// TIA Portal project "DistributoreCaffè" (V19)

(* hardware
DEVICE "S7-1200 station_1"  S7-1200 Station
   slot 0: "Telaio di montaggio_0"  S7-1200 Rack  Rack  V1.0
   slot 1: "PLC"  CPU 1212C DC/DC/Rly  6ES7 212-1HE40-0XB0  V4.6
DEVICE "HMI"  KTP900 Basic PN
   slot 0: "HMI_1"  KTP900 Basic PN  6AV2 123-2JB03-0AX0  17.0.0.0
   slot 1: "HMI_RT_1"  KTP900 Basic PN  6AV2 123-2JB03-0AX0  17.0.0.0
   slot 5: "HMI_1.IE_CP_1"  PROFINET Interface  17.0.0.0
      slot 1: "Interfaccia_1 PROFINET"  PROFINET Interface
         slot 1: "Porta_1"  Port
*)

// ===== PLC "PLC"  CPU 1212C DC/DC/Rly =====

TYPE "CreditoResto"
   STRUCT
      "5Cents" : Real;
      "10Cents" : Real;
      "20Cents" : Real;
      "50Cents" : Real;
      "1Euro" : Real;
      "2Euro" : Real;
   END_STRUCT;
END_TYPE

TYPE "RestoUtente"
   STRUCT
      "5Cents" : SInt;
      "10Cents" : SInt;
      "20Cents" : SInt;
      "50Cents" : SInt;
      "1Euro" : SInt;
      "2Euro" : SInt;
   END_STRUCT;
END_TYPE

TYPE "Prezzo"
   STRUCT
      Bevanda : String;
      Prezzo : Real;
   END_STRUCT;
END_TYPE

DATA_BLOCK "HMI"   // DB1
{ S7_Optimized_Access := 'TRUE' }
VERSION : 0.1
   VAR
      I5cents : Bool;
      I10Cents : Bool;
      I20Cents : Bool;
      I50Cents : Bool;
      I1Euro : Bool;
      I2Euro : Bool;
   END_VAR
   VAR RETAIN
      Resto : "RestoUtente";
   END_VAR
   VAR
      ValvolaBicchiere : Bool;
      ValvolaPaletta : Bool;
      ValvolaCaffè : Bool;
      ValvolaLatte : Bool;
      ValvolaGrappa : Bool;
      ValvolaZucchero : Bool;
      PrelievoProdotto : Bool;
   END_VAR
   VAR RETAIN
      ProdottoPronto : Bool;
   END_VAR
   VAR
      Corto : Bool;
      CortoMacchiato : Bool;
      CortoCorretto : Bool;
      CortoMacchiatoCorretto : Bool;
      Lungo : Bool;
      LungoMacchiato : Bool;
      LungoCorretto : Bool;
      LungoMacchiatoCorretto : Bool;
      ConfermaOrdine : Bool;
      BicchieriScarico : Bool;
      PaletteScarico : Bool;
      CaffèScarico : Bool;
      LatteScarico : Bool;
      GrappaScarico : Bool;
      ZuccheroScarico : Bool;
      Bicchieri : Int;
      Palette : Int;
      Caffè : SInt;
      Latte : SInt;
      Grappa : SInt;
      Zucchero : SInt;
      Credito : Real;
      Introiti : Real;
      PrelievoIntroiti : Bool;
      CreditoInsufficiente : Bool;
      QuantitàZuccheroSelezionata : SInt;
      RiduzioneZucchero : Bool;
      IncrementoZucchero : Bool;
      ProdottoInPreparazione : Bool;
   END_VAR
BEGIN
END_DATA_BLOCK

DATA_BLOCK "Sistema"   // DB2
{ S7_Optimized_Access := 'TRUE' }
VERSION : 0.1
   VAR RETAIN
      CreditoResto : "CreditoResto";
   END_VAR
   VAR
      PConfermaOrdine : Bool;
      BloccoInterfacciaUtente : Bool;
      NPrelievoProdotto : Bool;
      BevandaSelezionata : SInt;
      PCorto : Bool;
      PCortoMacchiato : Bool;
      PCortoCorretto : Bool;
      PCortoMacchiatoCorretto : Bool;
      PLungo : Bool;
      PLungoMacchiato : Bool;
      PLungoCorretto : Bool;
      PLungoMacchiatoCorretto : Bool;
      PPiùZucchero : Bool;
      PMenoZucchero : Bool;
   END_VAR
   VAR RETAIN
      Prezzi : Array[1..8] of "Prezzo";
   END_VAR
   VAR
      PBloccoInterfacciaUtente : Bool;
      NPrelievoProdotto2 : Bool;
   END_VAR
BEGIN
   CreditoResto."5Cents" := 5.0;
   CreditoResto."10Cents" := 5.0;
   CreditoResto."20Cents" := 5.0;
   CreditoResto."50Cents" := 5.0;
   CreditoResto."1Euro" := 5.0;
   CreditoResto."2Euro" := 5.0;
   Prezzi[1].Bevanda := 'Corto';
   Prezzi[1].Prezzo := 0.3;
   Prezzi[2].Bevanda := 'CortoMacchiato';
   Prezzi[2].Prezzo := 0.4;
   Prezzi[3].Bevanda := 'CortoCorretto';
   Prezzi[3].Prezzo := 0.4;
   Prezzi[4].Bevanda := 'CortoMacchiatoCorretto';
   Prezzi[4].Prezzo := 0.5;
   Prezzi[5].Bevanda := 'Lungo';
   Prezzi[5].Prezzo := 0.6;
   Prezzi[6].Bevanda := 'LungoMacchiato';
   Prezzi[6].Prezzo := 0.7;
   Prezzi[7].Bevanda := 'LungoCorretto';
   Prezzi[7].Prezzo := 0.7;
   Prezzi[8].Bevanda := 'LungoMacchiatoCorretto';
   Prezzi[8].Prezzo := 0.8;
END_DATA_BLOCK

DATA_BLOCK "AggiornamentoCreditoUtente_DB"   // DB3
{ S7_Optimized_Access := 'TRUE' }
VERSION : 0.1
// stored: InstanceOfName AggiornamentoCreditoUtenteCreditoDistributore
"AggiornamentoCreditoUtenteCreditoDistributore"
BEGIN
END_DATA_BLOCK

DATA_BLOCK "PreparazioneBevanda_DB"   // DB4
{ S7_Optimized_Access := 'TRUE' }
VERSION : 0.1
// stored: InstanceOfName PreparazioneBevanda
"PreparazioneBevanda"
BEGIN
END_DATA_BLOCK

DATA_BLOCK "AggiornamentoRestoUtenteCreditoUtenteCreditoDistributore_DB"   // DB5
{ S7_Optimized_Access := 'TRUE' }
VERSION : 0.1
// stored: InstanceOfName AggiornamentoRestoUtenteCreditoUtenteCreditoDistributore
"AggiornamentoRestoUtenteCreditoUtenteCreditoDistributore"
BEGIN
END_DATA_BLOCK

FUNCTION_BLOCK "AggiornamentoCreditoUtenteCreditoDistributore"   // FB1, LAD
{ S7_Optimized_Access := 'TRUE' }
VERSION : 0.1
   VAR_INPUT
      "5Cents" : Bool;
      "10Cents" : Bool;
      "20Cents" : Bool;
      "50Cents" : Bool;
      "1Euro" : Bool;
      "2Euro" : Bool;
   END_VAR
   VAR_IN_OUT
      CreditoDistributore : "CreditoResto";
      CreditoUtente : Real;
   END_VAR
   VAR
      PI5Cents : Bool;
      PI10Cents : Bool;
      PI20Cents : Bool;
      PI50Cents : Bool;
      PI1Euro : Bool;
      PI2Euro : Bool;
   END_VAR
   VAR_TEMP   // added for the SCL form of the ladder/FBD networks
      _w1 : Bool;
      _w2 : Bool;
      _w3 : Bool;
      _w4 : Bool;
      _w5 : Bool;
      _w6 : Bool;
   END_VAR
BEGIN

REGION Network 1
   // Attenzione: i valori Real non sempre vengono salvati a cifra tonda
   // (Es: 0.2999999999.. oppure 0.31111111.. invece di 0.3)
   // Arrotondare dopo ogni operazione matematica che li implica
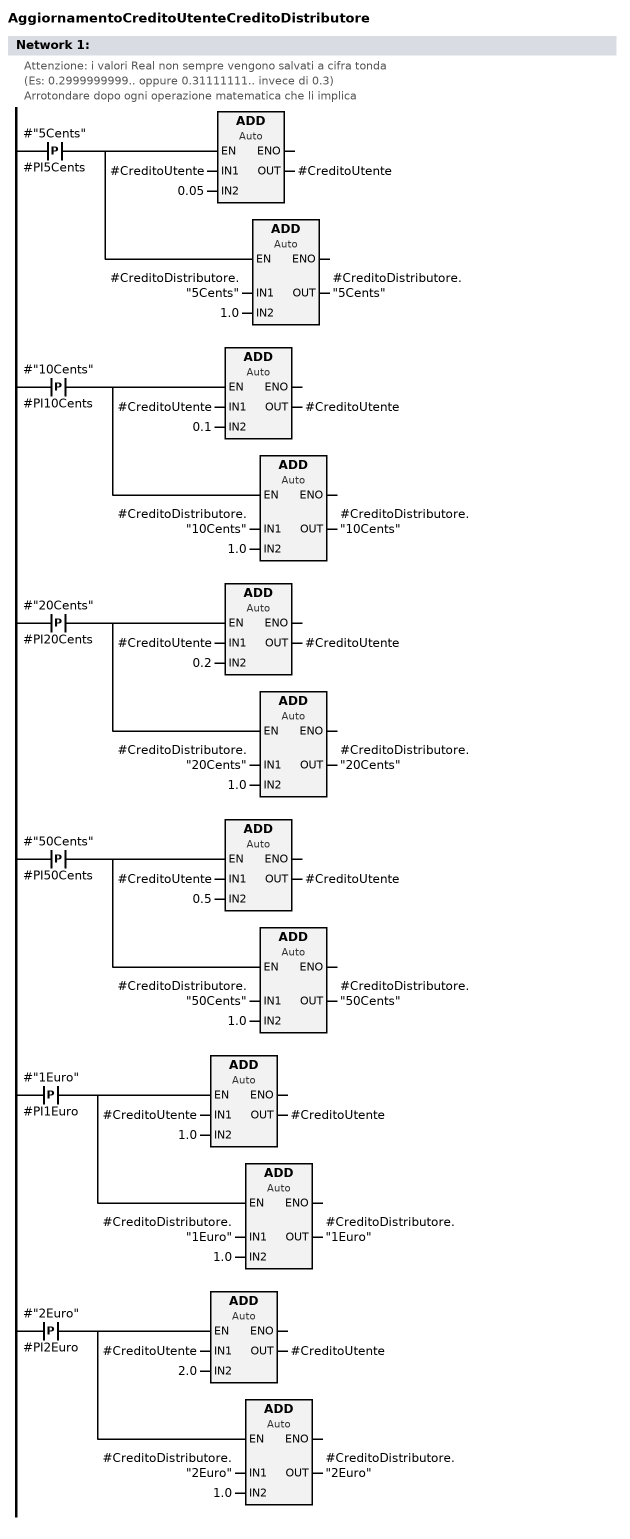
   RUNG wire#powerrail
      P_Contact(operand := #"5Cents", bit := #PI5Cents)
      wire#w1
      Add(in1 := #CreditoUtente, in2 := 0.05, out => #CreditoUtente)
   END_RUNG
   RUNG wire#w1
      Add(in1 := #CreditoDistributore."5Cents", in2 := 1.0, out => #CreditoDistributore."5Cents")
   END_RUNG
   RUNG wire#powerrail
      P_Contact(operand := #"10Cents", bit := #PI10Cents)
      wire#w2
      Add(in1 := #CreditoUtente, in2 := 0.1, out => #CreditoUtente)
   END_RUNG
   RUNG wire#w2
      Add(in1 := #CreditoDistributore."10Cents", in2 := 1.0, out => #CreditoDistributore."10Cents")
   END_RUNG
   RUNG wire#powerrail
      P_Contact(operand := #"20Cents", bit := #PI20Cents)
      wire#w3
      Add(in1 := #CreditoUtente, in2 := 0.2, out => #CreditoUtente)
   END_RUNG
   RUNG wire#w3
      Add(in1 := #CreditoDistributore."20Cents", in2 := 1.0, out => #CreditoDistributore."20Cents")
   END_RUNG
   RUNG wire#powerrail
      P_Contact(operand := #"50Cents", bit := #PI50Cents)
      wire#w4
      Add(in1 := #CreditoUtente, in2 := 0.5, out => #CreditoUtente)
   END_RUNG
   RUNG wire#w4
      Add(in1 := #CreditoDistributore."50Cents", in2 := 1.0, out => #CreditoDistributore."50Cents")
   END_RUNG
   RUNG wire#powerrail
      P_Contact(operand := #"1Euro", bit := #PI1Euro)
      wire#w5
      Add(in1 := #CreditoUtente, in2 := 1.0, out => #CreditoUtente)
   END_RUNG
   RUNG wire#w5
      Add(in1 := #CreditoDistributore."1Euro", in2 := 1.0, out => #CreditoDistributore."1Euro")
   END_RUNG
   RUNG wire#powerrail
      P_Contact(operand := #"2Euro", bit := #PI2Euro)
      wire#w6
      Add(in1 := #CreditoUtente, in2 := 2.0, out => #CreditoUtente)
   END_RUNG
   RUNG wire#w6
      Add(in1 := #CreditoDistributore."2Euro", in2 := 1.0, out => #CreditoDistributore."2Euro")
   END_RUNG
   // the same network as SCL:
   #_w1 := #"5Cents" AND NOT #PI5Cents;   // rising edge of #"5Cents"
   #PI5Cents := #"5Cents";
   IF #_w1 THEN
       #CreditoUtente := #CreditoUtente + 0.05;
       #CreditoDistributore."5Cents" := #CreditoDistributore."5Cents" + 1.0;
   END_IF;
   #_w2 := #"10Cents" AND NOT #PI10Cents;   // rising edge of #"10Cents"
   #PI10Cents := #"10Cents";
   IF #_w2 THEN
       #CreditoUtente := #CreditoUtente + 0.1;
       #CreditoDistributore."10Cents" := #CreditoDistributore."10Cents" + 1.0;
   END_IF;
   #_w3 := #"20Cents" AND NOT #PI20Cents;   // rising edge of #"20Cents"
   #PI20Cents := #"20Cents";
   IF #_w3 THEN
       #CreditoUtente := #CreditoUtente + 0.2;
       #CreditoDistributore."20Cents" := #CreditoDistributore."20Cents" + 1.0;
   END_IF;
   #_w4 := #"50Cents" AND NOT #PI50Cents;   // rising edge of #"50Cents"
   #PI50Cents := #"50Cents";
   IF #_w4 THEN
       #CreditoUtente := #CreditoUtente + 0.5;
       #CreditoDistributore."50Cents" := #CreditoDistributore."50Cents" + 1.0;
   END_IF;
   #_w5 := #"1Euro" AND NOT #PI1Euro;   // rising edge of #"1Euro"
   #PI1Euro := #"1Euro";
   IF #_w5 THEN
       #CreditoUtente := #CreditoUtente + 1.0;
       #CreditoDistributore."1Euro" := #CreditoDistributore."1Euro" + 1.0;
   END_IF;
   #_w6 := #"2Euro" AND NOT #PI2Euro;   // rising edge of #"2Euro"
   #PI2Euro := #"2Euro";
   IF #_w6 THEN
       #CreditoUtente := #CreditoUtente + 2.0;
       #CreditoDistributore."2Euro" := #CreditoDistributore."2Euro" + 1.0;
   END_IF;
END_REGION
END_FUNCTION_BLOCK

FUNCTION_BLOCK "PreparazioneBevanda"   // FB2, LAD
{ S7_Optimized_Access := 'TRUE' }
VERSION : 0.1
   VAR_INPUT
      BevandaSelezionata : SInt;
      InnescoProcesso : Bool;
   END_VAR
   VAR
      TPBicchiere : TP_TIME;
      NQTPBicchiere : Bool;
      TPPaletta : TP_TIME;
      NQTPPaletta : Bool;
      TPCaffè : TP_TIME;
      NQTPCaffè : Bool;
      TPLatte : TP_TIME;
      NQTPLatte : Bool;
      TPGrappa : TP_TIME;
      NQTPGrappa : Bool;
      TPzucchero : TP_TIME;
      NQTPZucchero : Bool;
      PInnescoProcesso : Bool;
   END_VAR
   VAR_TEMP
      PTZucchero : Int;
   END_VAR
   VAR_TEMP   // added for the SCL form of the ladder/FBD networks
      _w1 : Bool;
      _w2 : Bool;
      _w3 : Bool;
      _w4 : Bool;
      _w5 : Bool;
      _w6 : Bool;
      _w7 : Bool;
      _w8 : Bool;
      _w9 : Bool;
      _w10 : Bool;
      _w11 : Bool;
      _w12 : Bool;
   END_VAR
BEGIN

REGION Network 1
   // Gestire trigger timer valvole
   // - grappa caso bevanda corretta non macchiata
   // - zucchero caso bevanda zuccherata liscia o macchiata
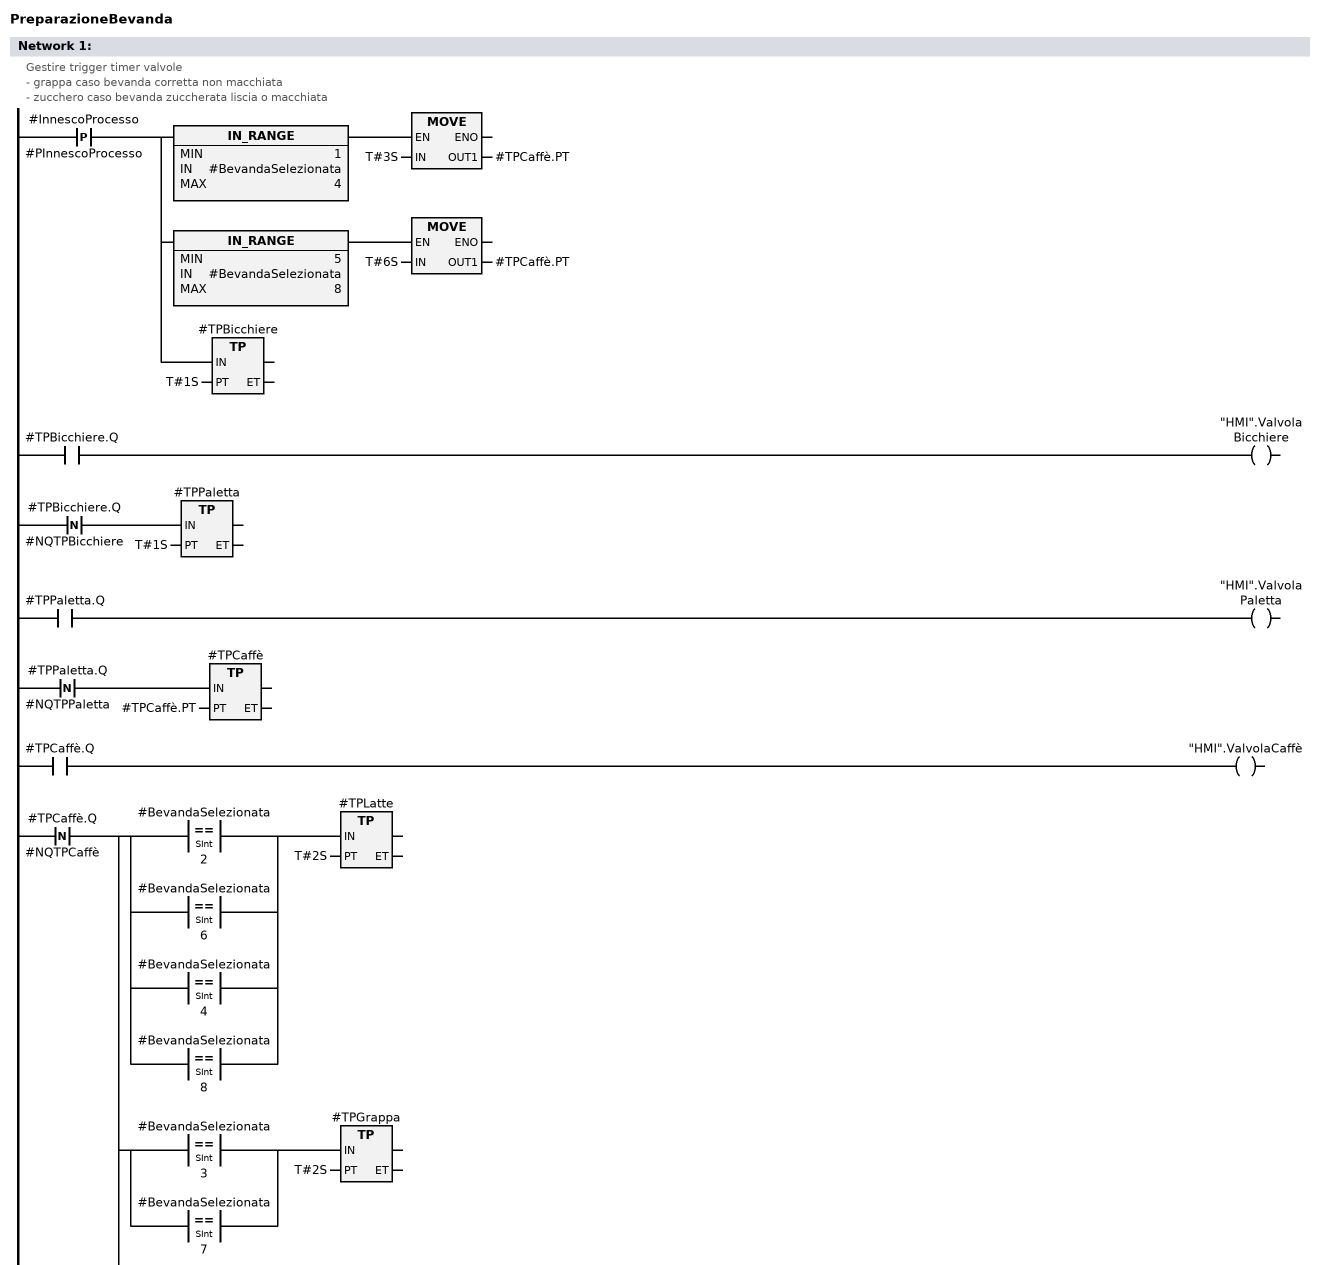
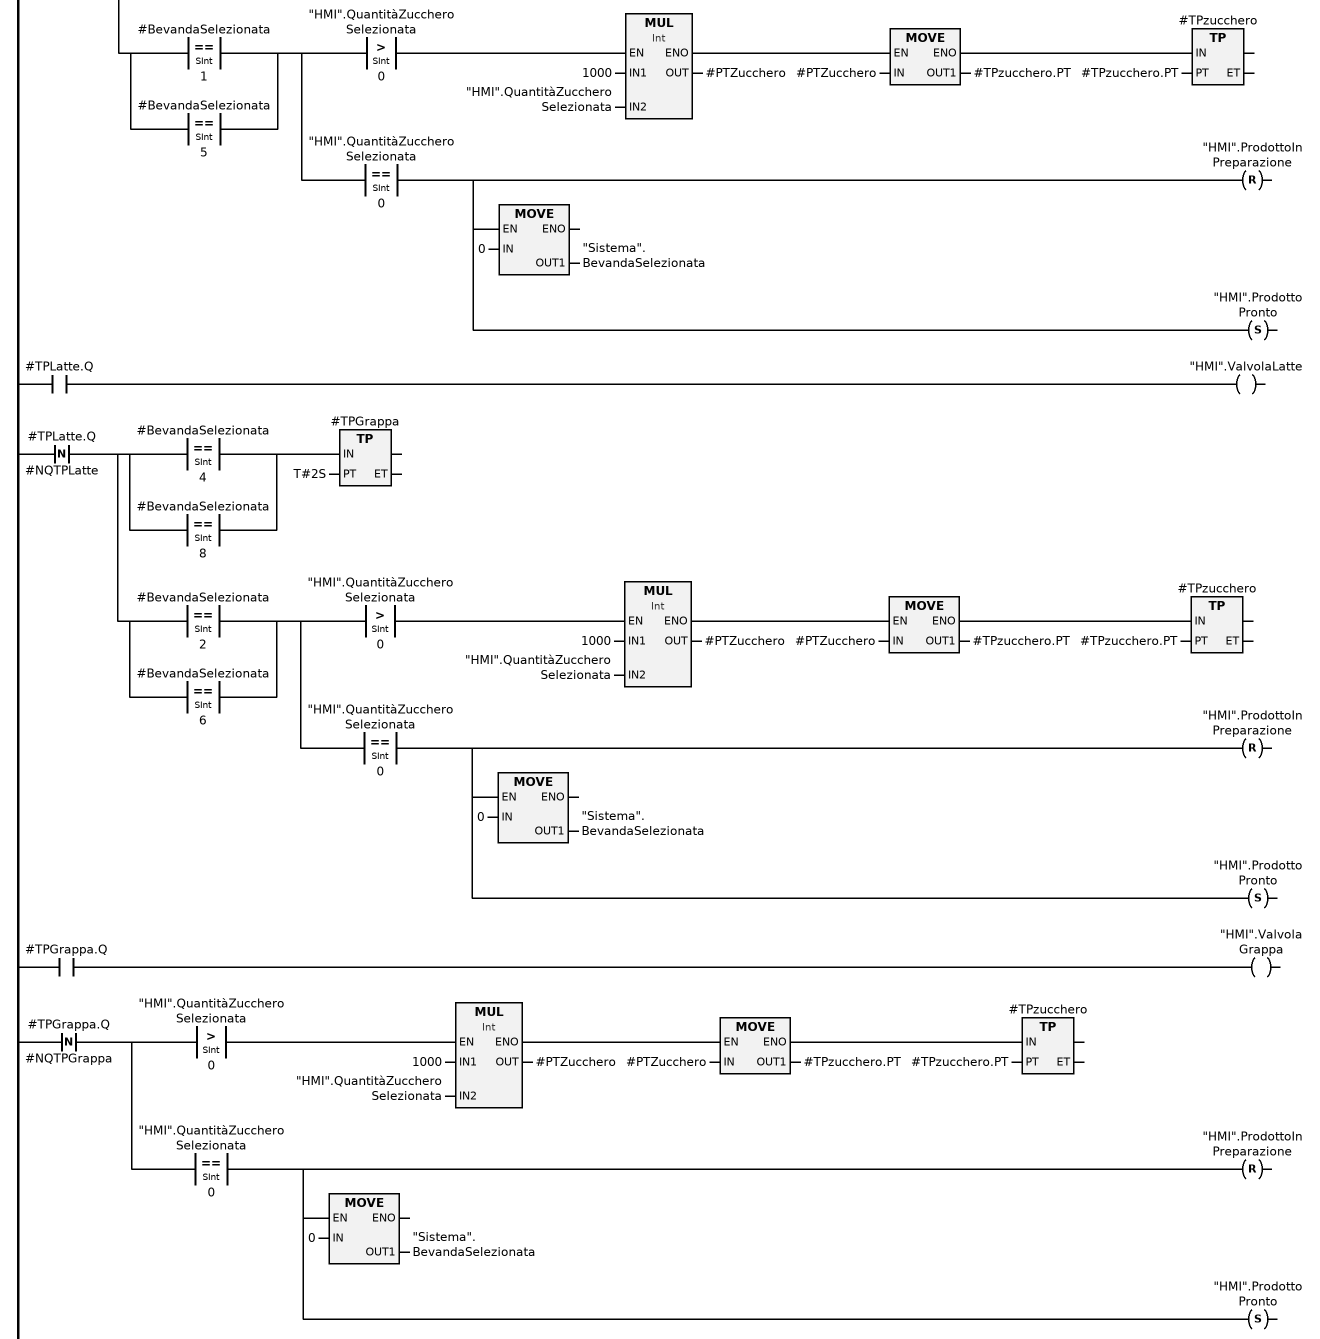
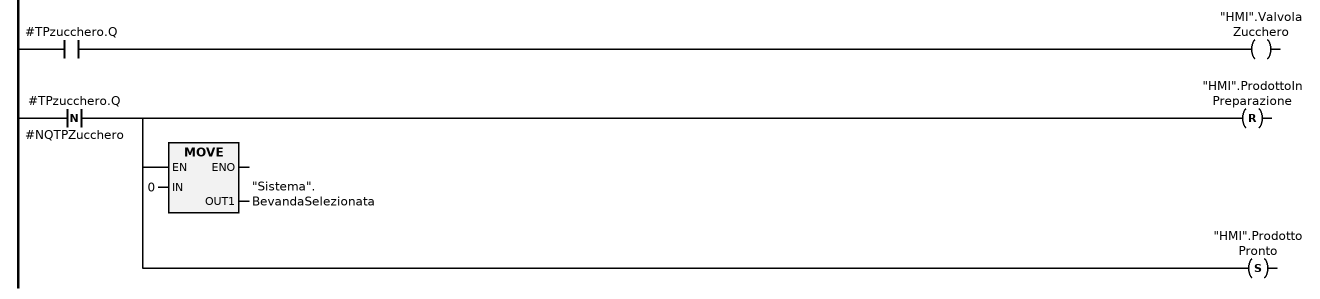
   #_w1 := #InnescoProcesso AND NOT #PInnescoProcesso;   // rising edge of #InnescoProcesso
   #PInnescoProcesso := #InnescoProcesso;
   IF #_w1 AND (1 <= #BevandaSelezionata) AND (#BevandaSelezionata <= 4) THEN #TPCaffè.PT := T#3S; END_IF;
   IF #_w1 AND (5 <= #BevandaSelezionata) AND (#BevandaSelezionata <= 8) THEN #TPCaffè.PT := T#6S; END_IF;
   #TPBicchiere(IN := #_w1, PT := T#1S);   // TP
   "HMI".ValvolaBicchiere := #TPBicchiere.Q;
   #_w2 := NOT #TPBicchiere.Q AND #NQTPBicchiere;   // falling edge of #TPBicchiere.Q
   #NQTPBicchiere := #TPBicchiere.Q;
   #TPPaletta(IN := #_w2, PT := T#1S);   // TP
   "HMI".ValvolaPaletta := #TPPaletta.Q;
   #_w3 := NOT #TPPaletta.Q AND #NQTPPaletta;   // falling edge of #TPPaletta.Q
   #NQTPPaletta := #TPPaletta.Q;
   #TPCaffè(IN := #_w3, PT := #TPCaffè.PT);   // TP
   "HMI".ValvolaCaffè := #TPCaffè.Q;
   #_w4 := NOT #TPCaffè.Q AND #NQTPCaffè;   // falling edge of #TPCaffè.Q
   #NQTPCaffè := #TPCaffè.Q;
   #TPLatte(IN := #_w4 AND ((#BevandaSelezionata = 2) OR (#BevandaSelezionata = 6) OR (#BevandaSelezionata = 4) OR (#BevandaSelezionata = 8)),   // TP
            PT := T#2S);
   #TPGrappa(IN := #_w4 AND ((#BevandaSelezionata = 3) OR (#BevandaSelezionata = 7)), PT := T#2S);   // TP
   #_w5 := #_w4 AND ((#BevandaSelezionata = 1) OR (#BevandaSelezionata = 5));
   #_w6 := #_w5 AND ("HMI".QuantitàZuccheroSelezionata > 0);
   IF #_w6 THEN
       #PTZucchero := 1000 * "HMI".QuantitàZuccheroSelezionata;
       #TPzucchero.PT := #PTZucchero;
   END_IF;
   #TPzucchero(IN := #_w6, PT := #TPzucchero.PT);   // TP
   IF #_w5 AND ("HMI".QuantitàZuccheroSelezionata = 0) THEN
       "HMI".ProdottoInPreparazione := FALSE;
       "Sistema".BevandaSelezionata := 0;
       "HMI".ProdottoPronto := TRUE;
   END_IF;
   "HMI".ValvolaLatte := #TPLatte.Q;
   #_w7 := NOT #TPLatte.Q AND #NQTPLatte;   // falling edge of #TPLatte.Q
   #NQTPLatte := #TPLatte.Q;
   #TPGrappa(IN := #_w7 AND ((#BevandaSelezionata = 4) OR (#BevandaSelezionata = 8)), PT := T#2S);   // TP
   #_w8 := #_w7 AND ((#BevandaSelezionata = 2) OR (#BevandaSelezionata = 6));
   #_w9 := #_w8 AND ("HMI".QuantitàZuccheroSelezionata > 0);
   IF #_w9 THEN
       #PTZucchero := 1000 * "HMI".QuantitàZuccheroSelezionata;
       #TPzucchero.PT := #PTZucchero;
   END_IF;
   #TPzucchero(IN := #_w9, PT := #TPzucchero.PT);   // TP
   IF #_w8 AND ("HMI".QuantitàZuccheroSelezionata = 0) THEN
       "HMI".ProdottoInPreparazione := FALSE;
       "Sistema".BevandaSelezionata := 0;
       "HMI".ProdottoPronto := TRUE;
   END_IF;
   "HMI".ValvolaGrappa := #TPGrappa.Q;
   #_w10 := NOT #TPGrappa.Q AND #NQTPGrappa;   // falling edge of #TPGrappa.Q
   #NQTPGrappa := #TPGrappa.Q;
   #_w11 := #_w10 AND ("HMI".QuantitàZuccheroSelezionata > 0);
   IF #_w11 THEN
       #PTZucchero := 1000 * "HMI".QuantitàZuccheroSelezionata;
       #TPzucchero.PT := #PTZucchero;
   END_IF;
   #TPzucchero(IN := #_w11, PT := #TPzucchero.PT);   // TP
   IF #_w10 AND ("HMI".QuantitàZuccheroSelezionata = 0) THEN
       "HMI".ProdottoInPreparazione := FALSE;
       "Sistema".BevandaSelezionata := 0;
       "HMI".ProdottoPronto := TRUE;
   END_IF;
   "HMI".ValvolaZucchero := #TPzucchero.Q;
   #_w12 := NOT #TPzucchero.Q AND #NQTPZucchero;   // falling edge of #TPzucchero.Q
   #NQTPZucchero := #TPzucchero.Q;
   IF #_w12 THEN
       "HMI".ProdottoInPreparazione := FALSE;
       "Sistema".BevandaSelezionata := 0;
       "HMI".ProdottoPronto := TRUE;
   END_IF;
END_REGION
END_FUNCTION_BLOCK

FUNCTION_BLOCK "AggiornamentoRestoUtenteCreditoUtenteCreditoDistributore"   // FB3, SCL
{ S7_Optimized_Access := 'TRUE' }
VERSION : 0.1
   VAR_INPUT
      BevandaSelezionata : SInt;
      InnescoProcesso : Bool;
   END_VAR
   VAR_IN_OUT
      Resto : "RestoUtente";
      CreditoDistributore : "CreditoResto";
      CreditoUtente : Real;
   END_VAR
   VAR
      Inception_R_TRIG_Instance : R_TRIG;
   END_VAR
BEGIN
   #Inception_R_TRIG_Instance(CLK:=#InnescoProcesso,
                              Q=>#Inception_R_TRIG_Instance.Q);

   IF #Inception_R_TRIG_Instance.Q THEN
       // Attenzione: i valori Real non sempre vengono salvati a cifra tonda
       // (Es: 0.2999999999.. oppure 0.31111111.. invece di 0.3)
       // Arrotondare dopo ogni operazione matematica che li implica
       #CreditoUtente := #CreditoUtente - "Sistema".Prezzi[#BevandaSelezionata].Prezzo;

       // Quantizzazione resto nei tagli di moneta disponibili nel salvadanaio del distributore
       // fino ad azzeramento credito utente residuo
       // Qualora il credito distributore sia insufficiente il credito utente residuo resta disponibile
       // per i prossimi acquisti
       WHILE #CreditoUtente >= 2.0 DO
           IF #CreditoDistributore."2Euro" > 0 THEN // (I tipi di monete inseriti dall'utenza sono già confluiti nel credito del distributore)
               // Rimuovere monete dal credito distributore...
               #CreditoDistributore."2Euro" := #CreditoDistributore."2Euro" - 1.0;
               // ... Aggiungerle al resto utente
               #Resto."2Euro" := #Resto."2Euro" + 1;
               // Aggiornare credito utente residuo
               #CreditoUtente := #CreditoUtente - 2.0;
           ELSIF #CreditoDistributore."1Euro" > 0 THEN
               // Rimuovere monete dal credito distributore...
               #CreditoDistributore."1Euro" := #CreditoDistributore."1Euro" - 1.0;
               // ... Aggiungerle al resto utente
               #Resto."1Euro" := #Resto."1Euro" + 1;
               // Aggiornare credito utente residuo
               #CreditoUtente := #CreditoUtente - 1.0;
           ELSIF #CreditoDistributore."50Cents" > 0 THEN
               #CreditoDistributore."50Cents" := #CreditoDistributore."50Cents" - 1.0;
               #Resto."50Cents" := #Resto."50Cents" + 1;
               #CreditoUtente := #CreditoUtente - 0.5;
           ELSIF #CreditoDistributore."20Cents" > 0 THEN
               #CreditoDistributore."20Cents" := #CreditoDistributore."20Cents" - 1.0;
               #Resto."20Cents" := #Resto."20Cents" + 1;
               #CreditoUtente := #CreditoUtente - 0.2;
           ELSIF #CreditoDistributore."10Cents" > 0 THEN
               #CreditoDistributore."10Cents" := #CreditoDistributore."10Cents" - 1.0;
               #Resto."10Cents" := #Resto."10Cents" + 1;
               #CreditoUtente := #CreditoUtente - 0.1;
           ELSIF #CreditoDistributore."5Cents" > 0 THEN
               #CreditoDistributore."5Cents" := #CreditoDistributore."5Cents" - 1.0;
               #Resto."5Cents" := #Resto."5Cents" + 1;
               #CreditoUtente := #CreditoUtente - 0.05;
           END_IF;
       END_WHILE;

       WHILE #CreditoUtente >= 1.0 DO
           IF #CreditoDistributore."1Euro" > 0 THEN
               #CreditoDistributore."1Euro" := #CreditoDistributore."1Euro" - 1.0;
               #Resto."1Euro" := #Resto."1Euro" + 1;
               #CreditoUtente := #CreditoUtente - 1.0;
           ELSIF #CreditoDistributore."50Cents" > 0 THEN
               #CreditoDistributore."50Cents" := #CreditoDistributore."50Cents" - 1.0;
               #Resto."50Cents" := #Resto."50Cents" + 1;
               #CreditoUtente := #CreditoUtente - 0.5;
           ELSIF #CreditoDistributore."20Cents" > 0 THEN
               #CreditoDistributore."20Cents" := #CreditoDistributore."20Cents" - 1.0;
               #Resto."20Cents" := #Resto."20Cents" + 1;
               #CreditoUtente := #CreditoUtente - 0.2;
           ELSIF #CreditoDistributore."10Cents" > 0 THEN
               #CreditoDistributore."10Cents" := #CreditoDistributore."10Cents" - 1.0;
               #Resto."10Cents" := #Resto."10Cents" + 1;
               #CreditoUtente := #CreditoUtente - 0.1;
           ELSIF #CreditoDistributore."5Cents" > 0 THEN
               #CreditoDistributore."5Cents" := #CreditoDistributore."5Cents" - 1.0;
               #Resto."5Cents" := #Resto."5Cents" + 1;
               #CreditoUtente := #CreditoUtente - 0.05;
           END_IF;
       END_WHILE;

       WHILE #CreditoUtente >= 0.5 DO
           IF #CreditoDistributore."50Cents" > 0 THEN
               #CreditoDistributore."50Cents" := #CreditoDistributore."50Cents" - 1.0;
               #Resto."50Cents" := #Resto."50Cents" + 1;
               #CreditoUtente := #CreditoUtente - 0.5;
           ELSIF #CreditoDistributore."20Cents" > 0 THEN
               #CreditoDistributore."20Cents" := #CreditoDistributore."20Cents" - 1.0;
               #Resto."20Cents" := #Resto."20Cents" + 1;
               #CreditoUtente := #CreditoUtente - 0.2;
           ELSIF #CreditoDistributore."10Cents" > 0 THEN
               #CreditoDistributore."10Cents" := #CreditoDistributore."10Cents" - 1.0;
               #Resto."10Cents" := #Resto."10Cents" + 1;
               #CreditoUtente := #CreditoUtente - 0.1;
           ELSIF #CreditoDistributore."5Cents" > 0 THEN
               #CreditoDistributore."5Cents" := #CreditoDistributore."5Cents" - 1.0;
               #Resto."5Cents" := #Resto."5Cents" + 1;
               #CreditoUtente := #CreditoUtente - 0.05;
           END_IF;
       END_WHILE;

       WHILE #CreditoUtente >= 0.2 DO
           IF #CreditoDistributore."20Cents" > 0 THEN
               #CreditoDistributore."20Cents" := #CreditoDistributore."20Cents" - 1.0;
               #Resto."20Cents" := #Resto."20Cents" + 1;
               #CreditoUtente := #CreditoUtente - 0.2;
           ELSIF #CreditoDistributore."10Cents" > 0 THEN
               #CreditoDistributore."10Cents" := #CreditoDistributore."10Cents" - 1.0;
               #Resto."10Cents" := #Resto."10Cents" + 1;
               #CreditoUtente := #CreditoUtente - 0.1;
           ELSIF #CreditoDistributore."5Cents" > 0 THEN
               #CreditoDistributore."5Cents" := #CreditoDistributore."5Cents" - 1.0;
               #Resto."5Cents" := #Resto."5Cents" + 1;
               #CreditoUtente := #CreditoUtente - 0.05;
           END_IF;
       END_WHILE;

       WHILE #CreditoUtente >= 0.1 DO
           IF #CreditoDistributore."10Cents" > 0 THEN
               #CreditoDistributore."10Cents" := #CreditoDistributore."10Cents" - 1.0;
               #Resto."10Cents" := #Resto."10Cents" + 1;
               #CreditoUtente := #CreditoUtente - 0.1;
           ELSIF #CreditoDistributore."5Cents" > 0 THEN
               #CreditoDistributore."5Cents" := #CreditoDistributore."5Cents" - 1.0;
               #Resto."5Cents" := #Resto."5Cents" + 1;
               #CreditoUtente := #CreditoUtente - 0.05;
           END_IF;
       END_WHILE;

       WHILE #CreditoUtente >= 0.05 DO
           IF #CreditoDistributore."5Cents" > 0 THEN
               #CreditoDistributore."5Cents" := #CreditoDistributore."5Cents" - 1.0;
               #Resto."5Cents" := #Resto."5Cents" + 1;
               #CreditoUtente := #CreditoUtente - 0.05;
           END_IF;
       END_WHILE;

       // Aggiornamento introiti proprietario
       "AggiornamentoIntroiti"(CreditoDistributore:="Sistema".CreditoResto,
                               Introiti:="HMI".Introiti);

   END_IF;
END_FUNCTION_BLOCK

FUNCTION "AggiornamentoIntroiti" : Void   // FC1, SCL
{ S7_Optimized_Access := 'TRUE' }
VERSION : 0.1
   VAR_INPUT
      CreditoDistributore : "CreditoResto";
   END_VAR
   VAR_IN_OUT
      Introiti : Real;
   END_VAR
   VAR CONSTANT
      CreditoIniziale : Real := 19.25;
   END_VAR
BEGIN
   // Il credito iniziale, destinato all'erogazione agevolata del resto, non costituisce guadagno per il proprietario

   // Attenzione: i valori Real non sempre vengono salvati a cifra tonda
   // (Es: 0.2999999999.. oppure 0.31111111.. invece di 0.3)
   // Arrotondare dopo ogni operazione matematica che li implica

   #Introiti := #CreditoDistributore."2Euro" * 2 + #CreditoDistributore."1Euro" + #CreditoDistributore."50Cents" * 0.5 + #CreditoDistributore."20Cents" * 0.2 + #CreditoDistributore."10Cents" * 0.1 + #CreditoDistributore."5Cents" * 0.05 - #CreditoIniziale;
END_FUNCTION

FUNCTION "ValutazioneInsufficienzaCredito" : Void   // FC2, SCL
{ S7_Optimized_Access := 'TRUE' }
VERSION : 0.1
   VAR_INPUT
      BevandaSelezionata : SInt;
      CreditoUtente : Real;
   END_VAR
   VAR_IN_OUT
      CreditoInsufficiente : Bool;
   END_VAR
BEGIN
   IF #CreditoUtente < ("Sistema".Prezzi[#BevandaSelezionata].Prezzo) THEN
       #CreditoInsufficiente := TRUE;
   ELSE
       #CreditoInsufficiente := FALSE;
   END_IF;
END_FUNCTION

ORGANIZATION_BLOCK "Main"   // OB1, LAD, ProgramCycle
TITLE = "Main Program Sweep (Cycle)"
{ S7_Optimized_Access := 'TRUE' }
VERSION : 0.1
   VAR_INPUT
      Initial_Call : Bool;   // Initial call of this OB
      Remanence : Bool;   // =True, if remanent data are available
   END_VAR
   VAR_TEMP   // added for the SCL form of the ladder/FBD networks
      _w1 : Bool;
      _w2 : Bool;
      _w3 : Bool;
      _w4 : Bool;
      _w5 : Bool;
      _w6 : Bool;
      _w7 : Bool;
      _w8 : Bool;
      _w9 : Bool;
   END_VAR
BEGIN

REGION Network 1